
   (* make sure L does not exceed the limits of a string *)
   #N := LIMIT(MN:=0,IN:=#L,MX:=254) - LEN("TEMP".STR1);
   IF #N <= 0 THEN
       (* truncate the string at length N *)
       IF #"M" = 1 THEN
           "TEMP".STR2 := RIGHT(IN:="TEMP".STR1,L:=#L);
       ELSE
           "TEMP".STR2 := LEFT(IN:="TEMP".STR1,L:=#L);
       END_IF;
   ELSIF #"M" = 1 THEN
       (* connect fill characters at the beginning *)
       #SX := "FILL"(C:=#C,L:=#N);
       "TEMP".STR2 := CONCAT(IN1:=#SX,IN2:="TEMP".STR1);
   ELSIF #"M" = 2 THEN
       (* center str beween fill characters *)
       (* for an uneven number of fill characters, there is one more at the end *)
       #SX := "FILL"(C:=#C,L:=WORD_TO_INT(SHR(IN:=INT_TO_WORD(#N+1),N:=1)));
       "TEMP".STR2 := CONCAT(IN1:="TEMP".STR1,IN2:=#SX);
       #SX := LEFT(IN:=#SX,L:=WORD_TO_INT(SHR(IN:=INT_TO_WORD(#N),N:=1)));
       "TEMP".STR2 := CONCAT(IN1:=#SX,IN2:="TEMP".STR2);
   ELSE
       (* connect fill characters at the end *)
       #SX := "FILL"(C:=#C,L:=#N);
       "TEMP".STR2 := CONCAT(IN1:="TEMP".STR1,IN2:=#SX);
   END_IF;

   #FIX := "TEMP".STR2;

   (* revision histroy
   hm  29. mar. 2008   rev 1.0
       original release

   *)
END_FUNCTION

FUNCTION "FLOAT_TO_REAL" : Real   // FC250, SCL
TITLE = FLOAT_TO_REAL
{ S7_Optimized_Access := 'FALSE' }
AUTHOR : hugo
FAMILY : STRINGS
NAME : FLT2REAL
VERSION : 1.3
// FLT_TO_REAL converts a string to a REAL.
// the function ignores all wrong characters.
// the comma can be , or .
// the exponent has to start with capital E or lowercase e .
// 
// uses: DEC_TO_INT [FC233]
//       RIGHT [FC32]
//       EXPN [FC78]
   VAR_INPUT
      FLT : String[254];
   END_VAR
   VAR_TEMP
      tFLT : String[20];
      _FLT AT tFLT : Struct
         length : Byte;
         act_length : Byte;
         str : Array[1..20] of Byte;
      END_STRUCT;
      pt : Int;   // pt : POINTER TO ARRAY[1..20] OF BYTE;
      i : Int;
      X : Byte;
      sign : Int;
      stop : Int;
      tmp : DInt;
      d : Int;
   END_VAR
BEGIN


   #sign := 1;

   #tFLT := #FLT;

   #pt := 1;    //ADR(FLT);
   #stop := BYTE_TO_INT(#_FLT.act_length);    //LEN(FLT);
   #tmp := 0;
   #d := 0;

   (* we first check for sign and exit if first number or dot is reached *)
   FOR #i := 1 TO #stop DO
       #X := #_FLT.str[#i];   //pt^[i];
       IF BYTE_TO_INT(#X) > 47 AND BYTE_TO_INT(#X) < 58 OR BYTE_TO_INT(#X) = 46 THEN
           EXIT;
       ELSIF BYTE_TO_INT(#X) = 45 THEN
           (* code 45 is sign *)
           #sign := -1;
       END_IF;
   END_FOR;

   (* now we scan numbers till end or dot or E is reached *)
   FOR #i := #i TO #stop DO
       #X := #_FLT.str[#i];   //pt^[i];
       IF BYTE_TO_INT(#X) = 44 OR BYTE_TO_INT(#X) = 46 OR BYTE_TO_INT(#X) = 69 OR BYTE_TO_INT(#X) = 101 THEN
           EXIT;
       (* calculate the value of the digit *)
       ELSIF BYTE_TO_INT(#X) > 47 AND BYTE_TO_INT(#X) < 58 THEN
           #tmp := #tmp * 10 + BYTE_TO_INT(#X) - 48;
       END_IF;
   END_FOR;

   (* process the portion after the comma if comma or dot is reached exit if exponent starts *)
   IF BYTE_TO_INT(#X) = 44 OR BYTE_TO_INT(#X) = 46 THEN
       FOR #i := #i + 1 TO #stop DO
           #X := #_FLT.str[#i];   //pt^[i];
           IF BYTE_TO_INT(#X) = 69 OR BYTE_TO_INT(#X) = 101 THEN
               EXIT;
           ELSIF BYTE_TO_INT(#X) > 47 AND BYTE_TO_INT(#X) < 58 THEN
               #tmp := #tmp * 10 + BYTE_TO_INT(#X) - 48;
               #d := #d - 1;
           END_IF;
       END_FOR;
   END_IF;

   (* process exponent if present *)
   IF BYTE_TO_INT(#X) = 69 OR BYTE_TO_INT(#X) = 101 THEN
       #d := #d + "DEC_TO_INT"(RIGHT(IN:=#tFLT,L:=#stop - #i));
   END_IF;

   #FLOAT_TO_REAL :=  "EXPN"(X:=10,N:=#d) * DINT_TO_REAL(#tmp * #sign);



   (* revision histroy
   hm  22. jun. 2008   rev 1.0
       original release

   hm  2. oct. 2008    rev 1.1
       fixed an error, characters 8 and 9 would not be converted

   hm  22. oct. 2008   rev 1.2
       last fix was not done correctly

   hm  23. oct. 2008   rev 1.3
       optimzed code
   *)
END_FUNCTION

FUNCTION "FSTRING_TO_BYTE" : Byte   // FC251, SCL
TITLE = FSTRING_TO_BYTE
{ S7_Optimized_Access := 'FALSE' }
AUTHOR : hugo
FAMILY : STRINGS
NAME : FSTR2BY
VERSION : 1.1
// FSTRING_TO_BYTE converts a formatted string into a byte.
// the string can be of the form 2#01010, 8#7234, 16#2AD3 and 1234
// 
// uses: EQ_STRNG [FC10]
//       LEFT [FC20]
//       BIN_TO_BYTE [FC220]
//       RIGHT [FC32]
//       LEN [FC21]
//       OCT_TO_BYTE [FC276]
//       HEX_TO_BYTE [FC256]
//       DEC_TO_BYTE [FC231]
//       CLEAN [FC228]
//       FIND [FC11] 
//       MID [FC26] 
//       DELETE [FC4]
   VAR_INPUT
      IN : String[254];
   END_VAR
   VAR_TEMP
      tIN : String[12];
   END_VAR
BEGIN


   #tIN := #IN;

   IF LEFT(IN:=#tIN,L:=2) S_COMP '2#' THEN
       (* we need to convert binary *)
       #FSTRING_TO_BYTE := "BIN_TO_BYTE"(RIGHT(IN:=#tIN,L:=LEN(#tIN) - 2));
   ELSIF LEFT(IN:=#tIN,L:=2) S_COMP '8#' THEN
       (* weneed to convert octals *)
       #FSTRING_TO_BYTE := "OCT_TO_BYTE"(RIGHT(IN:=#tIN,L:=LEN(#tIN) - 2));
   ELSIF LEFT(IN:=#tIN,L:=3) S_COMP '16#' THEN
       (* we need to convert hexadecimal *)
       #FSTRING_TO_BYTE := "HEX_TO_BYTE"(RIGHT(IN:=#tIN,L:=LEN(#tIN) - 3));
   ELSE
       (* we assume decimal representation *)
       #FSTRING_TO_BYTE := "DEC_TO_BYTE"("CLEAN"(IN:=#tIN,CX:='0123456789'));
   END_IF;


   (* revision histroy
   hm  18. jun. 2008   rev 1.0
       original release

   hm  20. sep. 2008   rev 1.1
       changed length of input string from 20 to 12
   *)
END_FUNCTION

FUNCTION "FSTRING_TO_DWORD" : DWord   // FC252, SCL
TITLE = FSTRING_TO_DWORD
{ S7_Optimized_Access := 'FALSE' }
AUTHOR : hugo
FAMILY : STRINGS
NAME : FSTR2DW
VERSION : 1.1
// FSTRING_TO_BYTE converts a formatted string into a byte.
// the string can be of the form 2#01010, 8#7234, 16#2AD3 and 1234
// 
// uses: EQ_STRNG [FC10]
//       LEFT [FC20]
//       BIN_TO_DWORD [FC221]
//       RIGHT [FC32]
//       LEN [FC21]
//       OCT_TO_DWORD [FC277]
//       HEX_TO_DWORD [FC257]
//       DEC_TO_DWORD [FC232]
//       CLEAN [FC228]
//       FIND [FC11] 
//       MID [FC26] 
//       DELETE [FC4]
   VAR_INPUT
      IN : String[254];
   END_VAR
   VAR_TEMP
      tIN : String[40];
   END_VAR
BEGIN


   #tIN := #IN;

   IF LEFT(IN:=#tIN,L:=2) S_COMP '2#' THEN
       (* we need to convert binary *)
       #FSTRING_TO_DWORD := "BIN_TO_DWORD"(RIGHT(IN:=#tIN,L:=LEN(#tIN) - 2));
   ELSIF LEFT(IN:=#tIN,L:=2) S_COMP '8#' THEN
       (* weneed to convert octals *)
       #FSTRING_TO_DWORD := "OCT_TO_DWORD"(RIGHT(IN:=#tIN,L:=LEN(#tIN) - 2));
   ELSIF LEFT(IN:=#tIN,L:=3) S_COMP '16#' THEN
       (* we need to convert hexadecimal *)
       #FSTRING_TO_DWORD := "HEX_TO_DWORD"(RIGHT(IN:=#tIN,L:=LEN(#tIN) - 3));
   ELSE
       (* we assume decimal representation *)
       #FSTRING_TO_DWORD := "DEC_TO_DWORD"("CLEAN"(IN:=#tIN,CX:='0123456789'));
   END_IF;


   (* revision histroy
   hm  18. jun. 2008   rev 1.0
       original release

   hm  20. sep. 2008   rev 1.1
       changed length of input dtring from 20 to 40


   *)
END_FUNCTION

FUNCTION "FSTRING_TO_MONTH" : Int   // FC253, SCL
TITLE = FSTRING_TO_MONTH
{ S7_Optimized_Access := 'FALSE' }
AUTHOR : hugo
FAMILY : STRINGS
NAME : FSTR2MON
VERSION : 1.2
// FSTRING_TO_MONTH converts a string into a month, the string can be a name for the month or a number.
// the function is language sensitve when LANG > 1 and checks for all languages when LANG = 0; 
// 
// uses: SETUP [DB1]
//       LANGUAGE [DB4]
//       STRNG_I [FC38]
//       EQ_STRNG [FC10]
//       TRIM [FC285]
//       FIND [FC11] 
//       REPLACE [FC31] 
//       CAPITALIZE [FC224]
//       TO_UPPER [FC284] 
//       LOWERCASE [FC273]
//       TO_LOWER [FC282]
   VAR_INPUT
      MTH : String[254];
      LANG : Int;
   END_VAR
   VAR_TEMP
      tMTH : String[20];
      lx : Int;
   END_VAR
BEGIN


   #tMTH := #MTH;

   IF #LANG = 0 THEN #lx := "LANGUAGE".DEFAULT; ELSE #lx := MIN(IN1:=#LANG, IN2:="LANGUAGE".LMAX); END_IF;
   #tMTH := "TRIM"(#tMTH);
   #tMTH := "CAPITALIZE"("LOWERCASE"(#tMTH));

   FOR #FSTRING_TO_MONTH := 1 TO 12 DO
       IF #tMTH S_COMP "LANGUAGE".MONTHS[#lx, #FSTRING_TO_MONTH] THEN RETURN; END_IF;
       IF #tMTH S_COMP "LANGUAGE".MONTHS3[#lx, #FSTRING_TO_MONTH] THEN RETURN; END_IF;
   END_FOR;

   (* since no name matched try to decode as integer *)
   #FSTRING_TO_MONTH := S_CONV(#tMTH);




   (* revision histroy
   hm  25. sep. 2008   rev 1.0
       original release

   hm  19. oct. 2008    rev 1.1
       changed language setup constants

   hm  25. oct. 2008   rev 1.2
       optimized code
   *)
END_FUNCTION

FUNCTION "FSTRING_TO_WEEK" : Byte   // FC254, SCL
TITLE = FSTRING_TO_WEEK
{ S7_Optimized_Access := 'FALSE' }
AUTHOR : hugo
FAMILY : STRINGS
NAME : FSTR2WEK
VERSION : 1.1
// FSTRING_TO_WEEK converts a list of weekdays into a byte where each bit represents a day of the week.
// bit 6 = mo, 0 = su;
// 
// uses: SETUP [DB1]
//       LANGUAGE [DB4]
//       FIND [FC11]
//       FSTRING_TO_WEEKDAY [FC255]
//       STRNG_I [FC38] 
//       EQ_STRNG [FC10] 
//       TRIM [FC285] 
//       REPLACE [FC31]
//       CAPITALIZE [FC224] 
//       TO_UPPER [FC284]
//       LOWERCASE [FC273] 
//       TO_LOWER [FC282]
//       MID [FC26]
//       RIGHT [FC32]
//       LEN [FC21]
   VAR_INPUT
      WEEK : String[254];
      LANG : Int;
   END_VAR
   VAR_TEMP
      tWEEK : String[60];
      pos : Int;
   END_VAR
BEGIN


   #tWEEK := #WEEK;

   #pos := FIND(IN1:=#tWEEK,IN2:=',');
   WHILE #pos > 0 DO
       #FSTRING_TO_WEEK := #FSTRING_TO_WEEK OR SHR(IN:=BYTE#128,N:="FSTRING_TO_WEEKDAY"(WDAY:=MID(IN:=#tWEEK, L:=#pos - 1,P:=1), LANG:=#LANG));
       #tWEEK := RIGHT(IN:=#tWEEK,L:=LEN(#tWEEK) - #pos);
       #pos := FIND(IN1:=#tWEEK,IN2:=',');
   END_WHILE;
   #FSTRING_TO_WEEK := #FSTRING_TO_WEEK OR SHR(IN:=BYTE#128,N:="FSTRING_TO_WEEKDAY"(WDAY:=#tWEEK, LANG:=#LANG)) AND BYTE#127;


   (* revision histroy
   hm  18. jun. 2008   rev 1.0
       original release

   hm  25. oct. 2008   rev 1.1
       using language defauls and input lang
   *)
END_FUNCTION

FUNCTION "FSTRING_TO_WEEKDAY" : Int   // FC255, SCL
TITLE = FSTRING_TO_WEEKDAY
{ S7_Optimized_Access := 'FALSE' }
AUTHOR : hugo
FAMILY : STRINGS
NAME : FSTR2WD
VERSION : 1.2
// FSTRING_TO_WEEKDAY converts a weekday string into an integer 1..7.
// 
// uses: SETUP [DB1]
//       LANGUAGE [DB4]
//       STRNG_I [FC38]
//       EQ_STRNG [FC10]
//       TRIM [FC285]
//       FIND [FC11] 
//       REPLACE [FC31] 
//       CAPITALIZE [FC224]
//       TO_UPPER [FC284] 
//       LOWERCASE [FC273]
//       TO_LOWER [FC282]
   VAR_INPUT
      WDAY : String[254];
      LANG : Int;
   END_VAR
   VAR_TEMP
      tWDAY : String[20];
      tmp : String[2];
      i : Int;
      ly : Int;
   END_VAR
BEGIN


   #tWDAY := #WDAY;

   IF #LANG = 0 THEN #ly := "LANGUAGE".DEFAULT; ELSE #ly := MIN(IN1:=#LANG, IN2:="LANGUAGE".LMAX); END_IF;
   (* tmp needs to be calculated first otherwise find can return wrong values *)
   #tmp := "TRIM"(#tWDAY);
   #tmp := "CAPITALIZE"("LOWERCASE"(#tmp));
   FOR #i := 1 TO 7 DO
       IF "LANGUAGE".WEEKDAYS2[#ly, #i] S_COMP #tmp THEN
           #FSTRING_TO_WEEKDAY := #i;
           RETURN;
       END_IF;
   END_FOR;
   #FSTRING_TO_WEEKDAY := S_CONV(#tWDAY);




   (* revision histroy
   hm  18. jun. 2008   rev 1.0
       original release

   hm  18. jul. 2008   rev 1.1
       changed nested call of left(trim()) for compatibility reasons

   hm  25. oct. 2008   rev 1.2
       using language constants
   *)
END_FUNCTION

FUNCTION "HEX_TO_BYTE" : Byte   // FC256, SCL
TITLE = HEX_TO_BYTE
{ S7_Optimized_Access := 'FALSE' }
AUTHOR : hugo
FAMILY : STRINGS
NAME : HEX2BY
VERSION : 1.1
// HEX_TO_BYTE converts a Hexadecimal string into a byte.
   VAR_INPUT
      HEX : String[254];
      _HEX AT HEX : Struct
         length : Byte;
         act_length : Byte;
         str : Array[1..5] of Byte;
      END_STRUCT;
   END_VAR
   VAR_TEMP
      pt : Int;   // pt : POINTER TO BYTE;
      i : Int;
      X : Byte;
      stop : Int;
   END_VAR
BEGIN


   #pt := 1;    //ADR(hex);
   #stop := BYTE_TO_INT(#_HEX.act_length);   //LEN(hex);
   FOR #i := 1 TO #stop DO
       (* read the first character and subtract 48 to get value in decimal 0 = 48 *)
       #X := #_HEX.str[#pt];
       (* calculate the value of the digit *)
       IF BYTE_TO_INT(#X) > 47 AND BYTE_TO_INT(#X) < 58 THEN
           #HEX_TO_BYTE := INT_TO_BYTE(BYTE_TO_INT(SHL(IN:=#HEX_TO_BYTE,N:=4)) + BYTE_TO_INT(#X) - 48);
       ELSIF BYTE_TO_INT(#X) > 64 AND BYTE_TO_INT(#X) < 71 THEN
           #HEX_TO_BYTE := INT_TO_BYTE(BYTE_TO_INT(SHL(IN:=#HEX_TO_BYTE,N:=4)) + BYTE_TO_INT(#X) - 55);
       ELSIF BYTE_TO_INT(#X) > 96 AND BYTE_TO_INT(#X) < 103 THEN
           #HEX_TO_BYTE := INT_TO_BYTE(BYTE_TO_INT(SHL(IN:=#HEX_TO_BYTE,N:=4)) + BYTE_TO_INT(#X) - 87);
       END_IF;
       #pt := #pt + 1;
   END_FOR;


   (* revision histroy
   hm  18. jun. 2008   rev 1.0
       original release

   hm  20. sep.2008    rev 1.1
       changed length of input string from 20 to 5

   *)
END_FUNCTION

FUNCTION "HEX_TO_DWORD" : DWord   // FC257, SCL
TITLE = HEX_TO_DWORD
{ S7_Optimized_Access := 'FALSE' }
AUTHOR : hugo
FAMILY : STRINGS
NAME : HEX2DW
VERSION : 1.4
// HEX_TO_DWORD converts a Hexadecimal string into a DWORD.
   VAR_INPUT
      Hex : String[254];
   END_VAR
   VAR_TEMP
      tHex : String[20];
      _Hex AT tHex : Struct
         length : Byte;
         act_length : Byte;
         str : Array[1..20] of Byte;
      END_STRUCT;
      pt : Int;   // pt : POINTER TO BYTE;
      i : Int;
      X : Byte;
      stop : Int;
   END_VAR
BEGIN


   #tHex := #Hex;

   #pt := 1;    //ADR(hex);
   #stop := BYTE_TO_INT(#_Hex.act_length);   //LEN(hex);
   FOR #i := 1 TO #stop DO
       (* read the first character and subtract 48 to get value in decimal 0 = 48 *)
       #X := #_Hex.str[#pt];
       (* calculate the value of the digit *)
       IF BYTE_TO_INT(#X) > 47 AND BYTE_TO_INT(#X) < 58 THEN
           #HEX_TO_DWORD := DINT_TO_DWORD(DWORD_TO_DINT(SHL(IN:=#HEX_TO_DWORD,N:=4)) + BYTE_TO_DINT(#X) - 48);
       ELSIF BYTE_TO_INT(#X) > 64 AND BYTE_TO_INT(#X) < 71 THEN
           #HEX_TO_DWORD := DINT_TO_DWORD(DWORD_TO_DINT(SHL(IN:=#HEX_TO_DWORD,N:=4)) + BYTE_TO_DINT(#X) - 55);
       ELSIF BYTE_TO_INT(#X) > 96 AND BYTE_TO_INT(#X) < 103 THEN
           #HEX_TO_DWORD := DINT_TO_DWORD(DWORD_TO_DINT(SHL(IN:=#HEX_TO_DWORD,N:=4)) + BYTE_TO_DINT(#X) - 87);
       END_IF;
       #pt := #pt + 1;
   END_FOR;

   (* revision histroy
   hm  2.10.2007       rev 1.0
       original release

   hm  19.11.2007      rev 1.1
       changed type of function from int to dword

   hm  4. mar 2008      rev 1.2
       added support for a..f and return 0 for invalid string

   hm  29. mar. 2008   rev 1.3
       changed STRING to STRING(8)

   hm  18. jun. 2008   rev 1.4
       changed input hex to STRING(20)
       function now ignores wrong characters
   *)
END_FUNCTION

FUNCTION "IS_ALNUM" : Bool   // FC258, SCL
TITLE = IS_ALNUM
{ S7_Optimized_Access := 'FALSE' }
AUTHOR : kurt
FAMILY : STRINGS
NAME : IS_ALNUM
VERSION : 1.1
// ISC_ALNUM testet ob in einem string nur Zahlen 0..9 vorkommen.
//  
// uses: SETUP [DB1]
//       ISC_ALPHA [FC267]
//       ISC_NUM [FC271]
   VAR_INPUT
      str : String[254];
      _str AT str : Struct
         length : Byte;
         act_length : Byte;
         str : Array[1..254] of Byte;
      END_STRUCT;
   END_VAR
   VAR_TEMP
      L : Int;
      pt : Int;   // POINTER TO BYTE;
      pos : Int;
   END_VAR
BEGIN


   #pt := 1;    //ADR(str);
   #L := BYTE_TO_INT(#_str.act_length);
   FOR #pos := 1 TO #L DO
     IF NOT ("ISC_ALPHA"(#_str.str[#pt]) OR "ISC_NUM"(#_str.str[#pt])) THEN
       #IS_ALNUM := FALSE;
       RETURN;
     END_IF;
         #pt := #pt + 1;
   END_FOR;
   #IS_ALNUM := #L > 0;


   (* revision history
   hm  29. feb 2008    rev 1.0
       original version

   hm  29. mar. 2008   rev 1.1
       changed STRING to STRING(STRING_LENGTH)
   *)
END_FUNCTION

FUNCTION "IS_ALPHA" : Bool   // FC259, SCL
TITLE = IS_ALPHA
{ S7_Optimized_Access := 'FALSE' }
AUTHOR : kurt
FAMILY : STRINGS
NAME : IS_ALPHA
VERSION : 1.1
// IS_ALPHA testet ob in einem string nur Zeichen a-z oder A - Z vorkommen.
// 
// uses: SETUP [DB1]
//       ISC_ALPHA [FC267]
   VAR_INPUT
      str : String[254];
      _str AT str : Struct
         length : Byte;
         act_length : Byte;
         str : Array[1..254] of Byte;
      END_STRUCT;
   END_VAR
   VAR_TEMP
      L : Int;
      pt : Int;   // POINTER TO BYTE;
      pos : Int;
   END_VAR
BEGIN


   #pt := 1;                            //ADR(str);
   #L := BYTE_TO_INT(#_str.act_length);  //LEN(str);
   FOR #pos := 1 TO #L DO
       IF NOT "ISC_ALPHA"(#_str.str[#pt]) THEN
           #IS_ALPHA := FALSE;
           RETURN;
       END_IF;
           #pt := #pt + 1;
   END_FOR;
   #IS_ALPHA := #L > 0;


   (* revision history
   hm  29. feb 2008    rev 1.0
       original version

   hm  29. mar. 2008   rev 1.1
       changed STRING to STRING(STRING_LENGTH)
   *)
END_FUNCTION

FUNCTION "IS_CC" : Bool   // FC260, SCL
TITLE = IS_CC
{ S7_Optimized_Access := 'FALSE' }
AUTHOR : Tobias
FAMILY : STRINGS
NAME : IS_CC
VERSION : 1.1
// ISC_CC testet ob ein string nur aus Zeichen des Strings CMP besteht.
// 
// uses: LEN [FC21]
//       FIND [FC11]
//       MID [FC26]
   VAR_INPUT
      str : String[254];
      cmp : String[254];
   END_VAR
   VAR_TEMP
      tstr : String[254];
      tcmp : String[254];
      L : Int;
      pos : Int;
   END_VAR
BEGIN


   #tstr := #str;
   #tcmp := #cmp;

   #L := LEN(#tstr);
   FOR #pos := 1 TO #L DO
       IF FIND(IN1:=#tcmp,IN2:=MID(IN:=#tstr,L:=1,P:=#pos)) = 0 THEN RETURN; END_IF;
   END_FOR;
   #IS_CC := #L > 0;



   (* revision history
   hm  19. mar 2008    rev 1.0
       original version

   hm  29. mar. 2008   rev 1.1
       changed STRING to STRING(STRING_LENGTH)
   *)
END_FUNCTION

FUNCTION "IS_CTRL" : Bool   // FC261, SCL
TITLE = IS_CTRL
{ S7_Optimized_Access := 'FALSE' }
AUTHOR : kurt
FAMILY : STRINGS
NAME : ISCTRL
VERSION : 1.1
// IS_CTRL testet ob in einem string nur Steuerzeichen (Char < 32) vorkommen.
// 
// uses: ISC_CTRL [FC268]
   VAR_INPUT
      str : String[254];
      _str AT str : Struct
         length : Byte;
         act_length : Byte;
         str : Array[1..254] of Byte;
      END_STRUCT;
   END_VAR
   VAR_TEMP
      L : Int;
      pt : Int;   // POINTER TO BYTE;
      pos : Int;
   END_VAR
BEGIN


   #pt := 1;                            //ADR(str);
   #L := BYTE_TO_INT(#_str.act_length);  //LEN(str);
   FOR #pos := 1 TO #L DO
       IF NOT ("ISC_CTRL"(#_str.str[#pt])) THEN
           #IS_CTRL := FALSE;
           RETURN;
       END_IF;
           #pt := #pt + 1;
   END_FOR;
   #IS_CTRL := #L > 0;


   (* revision history
   hm  29. feb. 2008   rev 1.0
       original version

   hm  29. mar. 2008   rev 1.1
       changed STRING to STRING(STRING_LENGTH)
   *)
END_FUNCTION

FUNCTION "IS_HEX" : Bool   // FC262, SCL
TITLE = IS_HEX
{ S7_Optimized_Access := 'FALSE' }
AUTHOR : kurt
FAMILY : STRINGS
NAME : ISHEX
VERSION : 1.1
// IS_HEX testet ob in einem string nur Zahlen 0..9 oder A..F oder a..f  vorkommen.
   VAR_INPUT
      str : String[254];
      _str AT str : Struct
         length : Byte;
         act_length : Byte;
         str : Array[1..254] of Byte;
      END_STRUCT;
   END_VAR
   VAR_TEMP
      L : Int;
      pt : Int;   // POINTER TO BYTE;
      pos : Int;
   END_VAR
BEGIN


   #pt := 1;                            //ADR(str);
   #L := BYTE_TO_INT(#_str.act_length);  //LEN(str);
   FOR #pos := 1 TO #L DO
       IF NOT ("ISC_HEX"(#_str.str[#pt])) THEN
           #IS_HEX := FALSE;
           RETURN;
       END_IF;
           #pt := #pt + 1;
   END_FOR;
   #IS_HEX := #L > 0;


   (* revision history
   hm  29. feb 2008    rev 1.0
       original version

   hm  29. mar. 2008   rev 1.1
       changed STRING to STRING(STRING_LENGTH)
   *)
END_FUNCTION

FUNCTION "IS_LOWER" : Bool   // FC263, SCL
TITLE = IS_LOWER
{ S7_Optimized_Access := 'FALSE' }
AUTHOR : kurt
FAMILY : STRINGS
NAME : ISLOWER
VERSION : 1.1
// IS_LOWER testet ob in einem string nur kleinbuchstaben vorkommen.
// 
// uses: SETUP [DB1]
//       ISC_LOWER [FC270]
   VAR_INPUT
      str : String[254];
      _str AT str : Struct
         length : Byte;
         act_length : Byte;
         str : Array[1..254] of Byte;
      END_STRUCT;
   END_VAR
   VAR_TEMP
      l : Int;
      pt : Int;   // POINTER TO BYTE;
      pos : Int;
   END_VAR
BEGIN


   #pt := 1;                            //ADR(str);
   #l := BYTE_TO_INT(#_str.act_length);  //LEN(str);
   FOR #pos := 1 TO #l DO
       IF NOT ("ISC_LOWER"(#_str.str[#pt])) THEN
           #IS_LOWER := FALSE;
           RETURN;
       END_IF;
           #pt := #pt + 1;
   END_FOR;
   #IS_LOWER := #l > 0;


   (* revision history
   hm  29. feb 2008    rev 1.0
       original version

   hm  29. mar. 2008   rev 1.1
       changed STRING to STRING(STRING_LENGTH)
   *)
END_FUNCTION

FUNCTION "IS_NCC" : Bool   // FC264, SCL
TITLE = IS_NCC
{ S7_Optimized_Access := 'FALSE' }
AUTHOR : Tobias
FAMILY : STRINGS
NAME : IS_NCC
VERSION : 1.1
// ISC_NCC testet ob in einem string keine Zeichen des Strings CMP enthalten sind.
//  
// uses: LEN [FC21]
//       FIND [FC11]
//       MID [FC26]
   VAR_INPUT
      str : String[254];
      cmp : String[254];
   END_VAR
   VAR_TEMP
      tstr : String[254];
      tcmp : String[254];
      L : Int;
      pos : Int;
   END_VAR
BEGIN


   #tstr := #str;
   #tcmp := #cmp;

   #L := LEN(#tstr);
   FOR #pos := 1 TO #L DO
       IF FIND(IN1:=#tcmp,IN2:=MID(IN:=#tstr,L:=1,P:=#pos)) > 0 THEN RETURN; END_IF;
   END_FOR;
   #IS_NCC := TRUE;



   (* revision history
   hm  19. mar 2008    rev 1.0
       original version

   hm  29. mar. 2008   rev 1.1
       changed STRING to STRING(STRING_LENGTH)
   *)
END_FUNCTION

FUNCTION "IS_NUM" : Bool   // FC265, SCL
TITLE = IS_NUM
{ S7_Optimized_Access := 'FALSE' }
AUTHOR : kurt
FAMILY : STRINGS
NAME : IS_NUM
VERSION : 1.1
// IS_NUM testet ob in einem string nur Zahlen 0..9 vorkommen.
//  
// uses: ISC_NUM [FC271]
   VAR_INPUT
      str : String[254];
      _str AT str : Struct
         length : Byte;
         act_length : Byte;
         str : Array[1..254] of Byte;
      END_STRUCT;
   END_VAR
   VAR_TEMP
      L : Int;
      pt : Int;   // POINTER TO BYTE;
      pos : Int;
   END_VAR
BEGIN


   #pt := 1;                            //ADR(str);
   #L := BYTE_TO_INT(#_str.act_length);  //LEN(str);
   FOR #pos := 1 TO #L DO
       IF NOT ("ISC_NUM"(#_str.str[#pt])) THEN
           #IS_NUM := FALSE;
           RETURN;
       END_IF;
           #pt := #pt + 1;
   END_FOR;
   #IS_NUM := #L > 0;


   (* revision history
   hm  29. feb 2008    rev 1.0
       original version

   hm  29. mar. 2008   rev 1.1
       changed STRING to STRING(STRING_LENGTH)
   *)
END_FUNCTION

FUNCTION "IS_UPPER" : Bool   // FC266, SCL
TITLE = IS_UPPER
{ S7_Optimized_Access := 'FALSE' }
AUTHOR : kurt
FAMILY : STRINGS
NAME : ISUPPER
VERSION : 1.1
// IS_UPPER testet ob in einem string keine Kleinbuchstaben vorkommen.
// 
// uses: SETUP [DB1]
//       ISC_UPPER [FC272]
   VAR_INPUT
      str : String[254];
      _str AT str : Struct
         length : Byte;
         act_length : Byte;
         str : Array[1..254] of Byte;
      END_STRUCT;
   END_VAR
   VAR_TEMP
      L : Int;
      pt : Int;   // POINTER TO BYTE;
      pos : Int;
   END_VAR
BEGIN


   #pt := 1;    //ADR(str);
   #L := BYTE_TO_INT(#_str.act_length);   //LEN(str);
   FOR #pos := 1 TO #L DO
       IF NOT ("ISC_UPPER"(#_str.str[#pt])) THEN
           #IS_UPPER := FALSE;
           RETURN;
       END_IF;
           #pt := #pt + 1;
   END_FOR;
   #IS_UPPER := #L > 0;


   (* revision history
   hm  29. feb 2008    rev 1.0
       original version

   hm  29. mar. 2008   rev 1.1
       changed STRING to STRING(STRING_LENGTH)
   *)
END_FUNCTION

FUNCTION "ISC_ALPHA" : Bool   // FC267, SCL
TITLE = ISC_ALPHA
{ S7_Optimized_Access := 'FALSE' }
AUTHOR : oscat
FAMILY : STRINGS
NAME : ISCALPHA
VERSION : 1.1
// ISC_ALPHA checks if a character is a..z or A..Z.
// 
// uses: SETUP [DB1]
   VAR_INPUT
      IN : Byte;
   END_VAR
BEGIN


   IF "SETUP".EXTENDED_ASCII THEN
       #ISC_ALPHA := (BYTE_TO_INT(#IN) > 64 AND BYTE_TO_INT(#IN) < 91) OR 
                    (BYTE_TO_INT(#IN) > 191  AND BYTE_TO_INT(#IN) <> 215 AND 
                     BYTE_TO_INT(#IN) <> 247) OR (BYTE_TO_INT(#IN) > 96 AND BYTE_TO_INT(#IN) < 123);
   ELSE
       #ISC_ALPHA := (BYTE_TO_INT(#IN) > 64 AND BYTE_TO_INT(#IN) < 91) OR 
                    (BYTE_TO_INT(#IN) > 96 AND BYTE_TO_INT(#IN) < 123);
   END_IF;

   (* revision history
   hm  6. mar. 2008    rev 1.0
       original version

   hm  19. oct. 2008   rev 1.1
       changes setup constants
   *)
END_FUNCTION

FUNCTION "ISC_CTRL" : Bool   // FC268, SCL
TITLE = ISC_CTRL
{ S7_Optimized_Access := 'FALSE' }
AUTHOR : oscat
FAMILY : STRINGS
NAME : ISC_CTRL
VERSION : 1.0
// ISC_ALPHA checks if a character is a control character.
   VAR_INPUT
      IN : Byte;
   END_VAR
BEGIN


   #ISC_CTRL := BYTE_TO_INT(#IN) < 32 OR BYTE_TO_INT(#IN) = 127;

   (* revision history
   hm    6. mar. 2008  rev 1.0
     original version

   *)
END_FUNCTION

FUNCTION "ISC_HEX" : Bool   // FC269, SCL
TITLE = ISC_HEX
{ S7_Optimized_Access := 'FALSE' }
AUTHOR : oscat
FAMILY : STRINGS
NAME : ISC_HEX
VERSION : 1.0
// ISC_HEX checks if a character is 0..9, A..F, a..f.
   VAR_INPUT
      IN : Byte;
   END_VAR
BEGIN


   #ISC_HEX := (BYTE_TO_INT(#IN) > 47 AND BYTE_TO_INT(#IN) < 58) OR (BYTE_TO_INT(#IN) > 64 AND BYTE_TO_INT(#IN) < 71) OR (BYTE_TO_INT(#IN) > 96 AND BYTE_TO_INT(#IN) < 103);

   (* revision history
   hm    6. mar. 2008  rev 1.0
     original version

   *)
END_FUNCTION

FUNCTION "ISC_LOWER" : Bool   // FC270, SCL
TITLE = ISC_LOWER
{ S7_Optimized_Access := 'FALSE' }
AUTHOR : hugo
FAMILY : STRINGS
NAME : ISCLOWER
VERSION : 1.1
// isc_lower checks if a character is lowercase.
// 
// uses: SETUP [DB1]
   VAR_INPUT
      IN : Byte;
   END_VAR
BEGIN


   IF "SETUP".EXTENDED_ASCII THEN
     #ISC_LOWER := ((BYTE_TO_INT(#IN) > 96) AND (BYTE_TO_INT(#IN) < 123)) OR ((BYTE_TO_INT(#IN) > 222) AND (BYTE_TO_INT(#IN) <> 247));
   ELSE
     #ISC_LOWER := ((BYTE_TO_INT(#IN) > 96) AND (BYTE_TO_INT(#IN) < 123));
   END_IF;

   (* revision history
   hm  6. mar. 2008  rev 1.0
       original version

   hm  19. oct. 2008   rev 1.1
       changes setup constants
   *)
END_FUNCTION

FUNCTION "ISC_NUM" : Bool   // FC271, SCL
TITLE = ISC_NUM
{ S7_Optimized_Access := 'FALSE' }
AUTHOR : oscat
FAMILY : STRINGS
NAME : ISC_NUM
VERSION : 1.0
// ISC_NUM checks if a character is 0..9.
   VAR_INPUT
      IN : Byte;
   END_VAR
BEGIN


   #ISC_NUM := BYTE_TO_INT(#IN) > 47 AND BYTE_TO_INT(#IN) < 58;

   (* revision history
   hm    6. mar. 2008  rev 1.0
     original version

   *)
END_FUNCTION

FUNCTION "ISC_UPPER" : Bool   // FC272, SCL
TITLE = ISC_UPPER
{ S7_Optimized_Access := 'FALSE' }
AUTHOR : hugo
FAMILY : STRINGS
NAME : ISCUPPER
VERSION : 1.1
// ISC_upper checks if a character is uppercase
// 
// uses: SETUP [DB1]
   VAR_INPUT
      IN : Byte;
   END_VAR
BEGIN


   IF "SETUP".EXTENDED_ASCII THEN
     #ISC_UPPER :=  ((BYTE_TO_INT(#IN) > 64) AND (BYTE_TO_INT(#IN) < 91)) OR (((BYTE_TO_INT(#IN) > 191) AND (BYTE_TO_INT(#IN) < 223)) AND (BYTE_TO_INT(#IN) <> 215));
   ELSE
     #ISC_UPPER := ((BYTE_TO_INT(#IN) > 64) AND (BYTE_TO_INT(#IN) < 91));
   END_IF;


   (* revision history
   hm  6. mar. 2008    rev 1.0
       original version

   hm  19. oct. 2008   rev 1.1
       changes setup constants

   *)
END_FUNCTION

